PopupScreen "RespirationRatios" 600x300
   TextField "Campo de texto_1" at 198,8 size 204x30; Text 'DATOS PACIENTE / PATIENT DATA'
   Button "Botón_6" at 429,255 size 146x32; TextOff 'Salida / Exit'
      on Click: function_efd93a16("RespirationRatios", 0, 0, 0, -1, 1)
   TextField "Campo de texto_4" at 31,88 size 123x29; Text 'Inspiración / Inspiration'
   IOField "Campo ES_1" at 159,86 size 110x35; FormatPattern 999.9; Unit %
      ProcessValue <- "OperatingParameters_InpirationRatio"
   TextField "Campo de texto_5" at 26,204 size 127x29; Text 'Esp+Retar / Esp+Delay'
   IOField "Campo ES_2" at 159,202 size 110x35; FormatPattern 999.9; Unit %
      ProcessValue <- "OperatingParameters_RestRatio"
   IOField "Campo ES_8" at 23,255 size 242x32; FormatPattern 99999999999999999999
      ProcessValue <- "DateTime_LocalDateOut"
   TextField "Campo de texto_6" at 33,126 size 121x29; Text 'Espiración / Espiration'
   IOField "Campo ES_3" at 159,124 size 110x35; FormatPattern 999.9; Unit %
      ProcessValue <- "OperatingParameters_EspirationRatio"
   TextField "Campo de texto_7" at 304,206 size 145x29; Text 'Rest. Tiempo / Rest. Time'
   TextField "Campo de texto_2" at 31,49 size 123x29; Text 'Frecuencia / Frequency'
   IOField "Campo ES_5" at 159,47 size 110x35; FormatPattern 99; Unit BPM
      ProcessValue <- "OperatingParameters_FrequencySetpoint"
   TextField "Campo de texto_3" at 300,51 size 148x29; Text 'Tiempo Ciclo / Cicle Time'
   IOField "Campo ES_6" at 453,49 size 110x35; FormatPattern 999999; Unit s
      ProcessValue <- "DataValues_TotalTime"
   TextField "Campo de texto_8" at 303,90 size 145x29; Text 'Tiempo Insp. / Insp. Time'
   IOField "Campo ES_7" at 453,88 size 110x35; FormatPattern 999999; Unit s
      ProcessValue <- "DataValues_InspirationTime"
   TextField "Campo de texto_9" at 297,128 size 151x29; Text 'Tiempo Esp. / Esp. Time'
   IOField "Campo ES_9" at 453,126 size 110x35; FormatPattern 999999; Unit s
      ProcessValue <- "DataValues_EspirationTime"
   TextField "Campo de texto_10" at 34,165 size 121x29; Text 'Retardo / Delay'
   IOField "Campo ES_10" at 160,163 size 110x35; FormatPattern 999.9; Unit %
      ProcessValue <- "OperatingParameters_DelayRatio"
   TextField "Campo de texto_11" at 269,167 size 180x29; Text 'Tiempo Retardo / Delay Time'
   IOField "Campo ES_11" at 454,165 size 110x35; FormatPattern 999999; Unit s
      ProcessValue <- "DataValues_DelayTime"
   IOField "Campo ES_4" at 453,204 size 110x35; FormatPattern 999999; Unit s
      ProcessValue <- "DataValues_RestTime"

screen "Graphics" 800x480
   Button "Botón_2" at 4,442 size 120x35; TextOff 'PARAMETROS / PARAMETERS'
      on Press: ActivateScreen("Parameters", 0)
   TextField "Campo de texto_2" at 9,163 size 69x25; Text 'Peep P'
   TextField "Campo de texto_1" at 8,41 size 53x25; Text 'Pip P'
   Button "Botón_35" at 11,235 size 48x39; TextOff '-'
      on Press: function_b14e0dd5("OperatingParameters_PeepPBMinus", 0)
      Visibility <- "AlwaysTRUE"
   Button "Botón_7" at 67,235 size 48x39; TextOff '+'
      on Press: function_b14e0dd5("OperatingParameters_PeepPBPlus", 0)
      Visibility <- "AlwaysTRUE"
   Button "Botón_4" at 10,113 size 48x39; TextOff '-'
      on Press: function_b14e0dd5("OperatingParameters_PeakPBMinus", 0)
      Visibility <- "AlwaysTRUE"
   Button "Botón_5" at 66,113 size 48x39; TextOff '+'
      on Press: function_b14e0dd5("OperatingParameters_PeakPBPlus", 0)
      Visibility <- "AlwaysTRUE"
   TextField "Campo de texto_3" at 10,283 size 29x25; Text 'FR'
   Button "Botón_1" at 11,356 size 48x39; TextOff '-'
      on Press: function_b14e0dd5("OperatingParameters_FrPBMinus", 0)
      Visibility <- "AlwaysTRUE"
   Button "Botón_6" at 67,356 size 48x39; TextOff '+'
      on Press: function_b14e0dd5("OperatingParameters_FrPBPlus", 0)
      Visibility <- "AlwaysTRUE"
   IOField "Campo ES_30" at 10,187 size 105x45; FormatPattern 999
      ProcessValue <- "OperatingParameters_PeepSetpoint"
   IOField "Campo ES_2" at 11,307 size 105x45; FormatPattern 999
      ProcessValue <- "OperatingParameters_FrequencySetpoint"
   IOField "Campo ES_4" at 10,66 size 105x45; FormatPattern 999
      ProcessValue <- "OperatingParameters_PipSetpoint"
   Button "Botón_13" at 4,404 size 120x35; TextOff 'MODO / MODE'; TextList "ModeSelected"
      on Press: function_efd93a16("ControlMode", 0, 0, -1, -1, 1)
      ProcessValue <- "OperatingParameters_ControlMode"
   IOField "Campo ES_6" at 3,2 size 120x35; FormatPattern 99999999999999999999
      ProcessValue <- "DateTime_LocalDateOut"
   Button "Botón_3" at 742,143 size 53x35; TextOff 'Trigger'
      Visibility <- "Clock_1Hz"
   Button "Botón_9" at 127,143 size 134x35; TextOff 'RECLUTAMIENTO ON / RECRUITMENT ON'
      on Press: function_b14e0dd5("OperatingParameters_RecruitmentOn", 0)
   Button "Botón_10" at 394,143 size 134x35; TextOff 'RECLUTAMIENTO OFF / RECRUITMENT OFF'
      on Press: function_b14e0dd5("OperatingParameters_RecruitmentOff", 0)
   IOField "Campo ES_5" at 302,143 size 89x35; FormatPattern 9999999
      ProcessValue <- "OperatingParameters_RecruitmentElap"
   GraphicView "Visor de gráficos_2" at 264,144 size 35x35; Picture "weather_warning_signal_alert_exclamation_icon_124159"
      Visibility <- "OperatingParameters_RecruitmentEnding"
   Button "Botón_12" at 532,143 size 61x35; TextOff 'Hr'
      Visibility <- "Clock_1Hz"
   Button "Botón_14" at 603,143 size 61x35; TextOff 'Aire / Air'
      Visibility <- "Clock_1Hz"
   Button "Botón_15" at 673,143 size 61x35; TextOff 'O2'
      Visibility <- "Clock_1Hz"
   Button "Botón_11" at 3,3 size 35x35; TextOff 'M'
      on Press: ActivateScreen("Start", 0)
   Button "Botón_8" at 92,2 size 35x35; TextOff 'M'
      on Press: ActivateScreen("Motor", 0)
   GraphicView "Visor de gráficos_1" at 264,144 size 35x35; Picture "Protective_Equipment-20-512"
      Visibility <- "OperatingParameters_RecruitmentRunning"
   IOField "Campo ES_14" at 130,442 size 70x35; FormatPattern 999
      ProcessValue <- "DataValues_PipValue"
   TextField "Campo de texto_5" at 145,418 size 35x25; Text 'Pip'
   IOField "Campo ES_11" at 485,442 size 70x35; FormatPattern 999
      ProcessValue <- "DataValues_TidalVolumeValue"
   TextField "Campo de texto_4" at 486,420 size 69x25; Text 'V.Tidal / Tidal V'
   IOField "Campo ES_1" at 272,442 size 70x35; FormatPattern 999
      ProcessValue <- "DataValues_PeepValue"
   TextField "Campo de texto_6" at 282,418 size 51x25; Text 'Peep'
   IOField "Campo ES_3" at 414,442 size 70x35; FormatPattern 999
      ProcessValue <- "DataValues_FrequencyValue"
   TextField "Campo de texto_7" at 435,419 size 29x25; Text 'FR'
   IOField "Campo ES_7" at 343,442 size 70x35; FormatPattern 999
      ProcessValue <- "DataValues_DrivingPressure"
   TextField "Campo de texto_8" at 344,419 size 68x25; Text 'Driv. P'
   IOField "Campo ES_8" at 201,442 size 70x35; Authorization "Operación"; FormatPattern 999
      ProcessValue <- "DataValues_PlateauValue"
   TextField "Campo de texto_9" at 196,418 size 76x25; Text 'Plateau'
   IOField "Campo ES_29" at 627,442 size 70x35; FormatPattern 999
      ProcessValue <- "OperatingParameters_TriggerSetpoint"
   TextField "Campo de texto_10" at 633,419 size 73x25; Text 'Trigger'
   IOField "Campo ES_23" at 556,442 size 70x35; FormatPattern 999
      ProcessValue <- "DataValues_MinumValue"
   TextField "Campo de texto_11" at 555,420 size 77x25; Text 'V Minut'
   Switch "Interruptor_1" at 708,421 size 91x56; TextOn 'ON'; CaptionText 'Operación / Operation'; TextOff 'OFF'
      ProcessValue <- "Operation_Operation_ON"
   Rectangle "Rectángulo_1" at 130,439 size 70x7
      Visibility <- "AlarmsRaw_PipDisplayAlarmHI"
   Rectangle "Rectángulo_5" at 130,439 size 70x7
      Visibility <- "AlarmsRaw_PipDisplayPreAlarmHI"
   Rectangle "Rectángulo_6" at 130,473 size 70x7
      Visibility <- "AlarmsRaw_PipDisplayAlarmLOW"
   Rectangle "Rectángulo_7" at 130,473 size 70x7
      Visibility <- "AlarmsRaw_PipDisplayPreAlarmLOW"
   Rectangle "Rectángulo_8" at 201,439 size 70x7
      Visibility <- "AlarmsRaw_PlateauDisplayAlarmHI"
   Rectangle "Rectángulo_9" at 201,439 size 70x7
      Visibility <- "AlarmsRaw_PlateauDisplayPreAlarmHI"
   Rectangle "Rectángulo_10" at 201,473 size 70x7
      Visibility <- "AlarmsRaw_PlateauDisplayAlarmHI"
   Rectangle "Rectángulo_11" at 201,473 size 70x7
      Visibility <- "AlarmsRaw_PlateauDisplayPreAlarmLOW"
   Rectangle "Rectángulo_12" at 272,439 size 70x7
      Visibility <- "AlarmsRaw_PeepDisplayAlarmHI"
   Rectangle "Rectángulo_13" at 272,439 size 70x7
      Visibility <- "AlarmsRaw_PeepDisplayPreAlarmHI"
   Rectangle "Rectángulo_14" at 272,472 size 70x7
      Visibility <- "AlarmsRaw_PeepDisplayAlarmLOW"
   Rectangle "Rectángulo_15" at 272,472 size 70x7
      Visibility <- "AlarmsRaw_PeepDisplayPreAlarmLOW"
   Rectangle "Rectángulo_16" at 343,439 size 70x7
      Visibility <- "AlarmsRaw_FrequencyDisplayAlarmHI"
   Rectangle "Rectángulo_17" at 343,439 size 70x7
      Visibility <- "AlarmsRaw_FrequencyDisplayPreAlarmHI"
   Rectangle "Rectángulo_18" at 343,472 size 70x7
      Visibility <- "AlarmsRaw_FrequencyDisplayAlarmLOW"
   Rectangle "Rectángulo_19" at 343,472 size 70x7
      Visibility <- "AlarmsRaw_FrequencyDisplayPreAlarmLOW"
   Rectangle "Rectángulo_20" at 414,439 size 70x7
      Visibility <- "AlarmsRaw_FrequencyDisplayAlarmHI"
   Rectangle "Rectángulo_21" at 414,439 size 70x7
      Visibility <- "AlarmsRaw_FrequencyDisplayPreAlarmHI"
   Rectangle "Rectángulo_22" at 414,472 size 70x7
      Visibility <- "AlarmsRaw_FrequencyDisplayAlarmLOW"
   Rectangle "Rectángulo_23" at 414,472 size 70x7
      Visibility <- "AlarmsRaw_FrequencyDisplayPreAlarmLOW"
   Rectangle "Rectángulo_24" at 485,439 size 70x7
      Visibility <- "AlarmsRaw_TidalVolumeDisplayAlarmHI"
   Rectangle "Rectángulo_25" at 485,439 size 70x7
      Visibility <- "AlarmsRaw_TidalVolumeDisplayPreAlarmHI"
   Rectangle "Rectángulo_26" at 485,472 size 70x7
      Visibility <- "AlarmsRaw_TidalVolumeDisplayAlarmLOW"
   Rectangle "Rectángulo_27" at 485,472 size 70x7
      Visibility <- "AlarmsRaw_TidalVolumeDisplayPreAlarmLOW"
   Rectangle "Rectángulo_28" at 556,439 size 70x7
      Visibility <- "AlarmsRaw_VolumeMinuteDisplayAlarmHI"
   Rectangle "Rectángulo_29" at 556,439 size 70x7
      Visibility <- "AlarmsRaw_VolumeMinuteDisplayPreAlarmHI"
   Rectangle "Rectángulo_30" at 556,472 size 70x7
      Visibility <- "AlarmsRaw_VolumeMinuteDisplayAlarmLOW"
   Rectangle "Rectángulo_31" at 556,472 size 70x7
      Visibility <- "AlarmsRaw_VolumeMinuteDisplayPreAlarmLOW"
   Rectangle "Rectángulo_32" at 627,439 size 70x7
      Visibility <- "AlarmsRaw_TriggerDisplayAlarmHI"
   Rectangle "Rectángulo_33" at 627,439 size 70x7
      Visibility <- "AlarmsRaw_TriggerDisplayPreAlarmHI"
   Rectangle "Rectángulo_34" at 627,472 size 70x7
      Visibility <- "AlarmsRaw_TriggerDisplayAlarmLOW"
   Rectangle "Rectángulo_35" at 627,472 size 70x7
      Visibility <- "AlarmsRaw_TriggerDisplayPreAlarmLOW"
   TrendView "Visor de curvas_2" at 127,182 size 669x239
   TrendView "Visor de curvas_1" at 126,2 size 669x137
*)